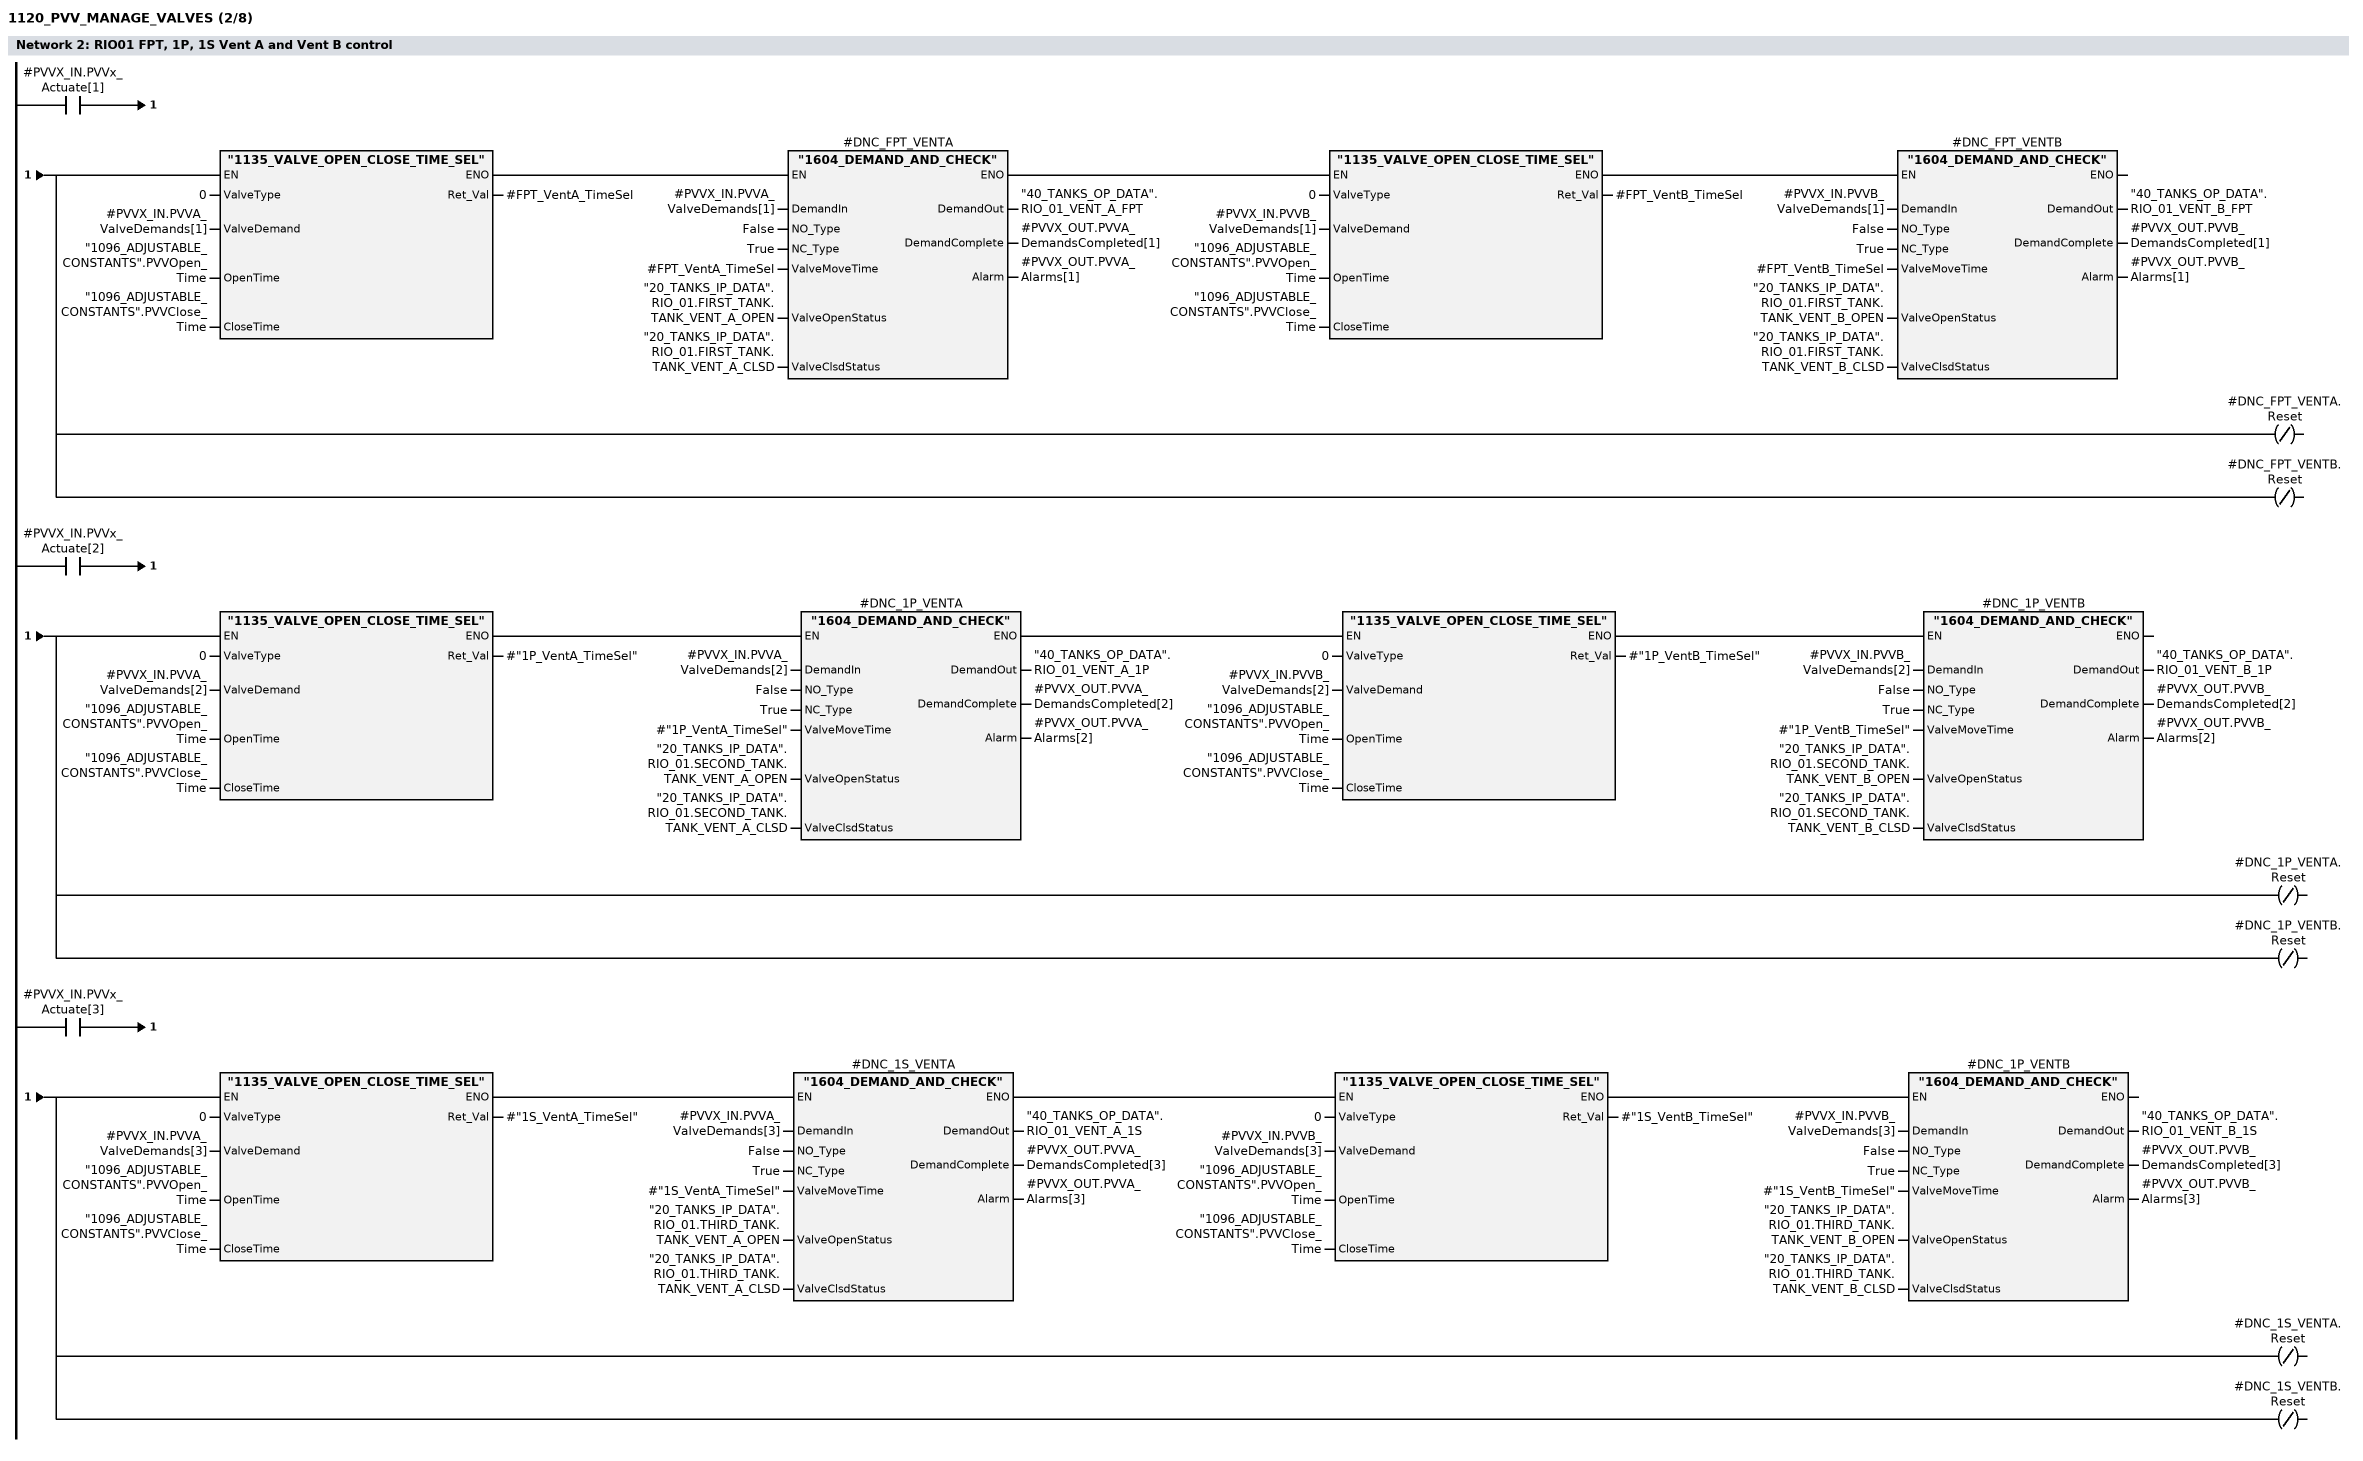
   RUNG wire#powerrail
      Contact( #PVVX_IN.PVVx_Actuate[1] )
      wire#w1
      "1135_VALVE_OPEN_CLOSE_TIME_SEL"(ValveType := 0, ValveDemand := #PVVX_IN.PVVA_ValveDemands[1], OpenTime := "1096_ADJUSTABLE_CONSTANTS".PVVOpen_Time, CloseTime := "1096_ADJUSTABLE_CONSTANTS".PVVClose_Time, Ret_Val => #FPT_VentA_TimeSel)
      #DNC_FPT_VENTA(DemandIn := #PVVX_IN.PVVA_ValveDemands[1], NO_Type := False, NC_Type := True, ValveMoveTime := #FPT_VentA_TimeSel, ValveOpenStatus := "20_TANKS_IP_DATA".RIO_01.FIRST_TANK.TANK_VENT_A_OPEN, ValveClsdStatus := "20_TANKS_IP_DATA".RIO_01.FIRST_TANK.TANK_VENT_A_CLSD, DemandOut => "40_TANKS_OP_DATA".RIO_01_VENT_A_FPT, DemandComplete => #PVVX_OUT.PVVA_DemandsCompleted[1], Alarm => #PVVX_OUT.PVVA_Alarms[1])
      "1135_VALVE_OPEN_CLOSE_TIME_SEL"(ValveType := 0, ValveDemand := #PVVX_IN.PVVB_ValveDemands[1], OpenTime := "1096_ADJUSTABLE_CONSTANTS".PVVOpen_Time, CloseTime := "1096_ADJUSTABLE_CONSTANTS".PVVClose_Time, Ret_Val => #FPT_VentB_TimeSel)
      #DNC_FPT_VENTB(DemandIn := #PVVX_IN.PVVB_ValveDemands[1], NO_Type := False, NC_Type := True, ValveMoveTime := #FPT_VentB_TimeSel, ValveOpenStatus := "20_TANKS_IP_DATA".RIO_01.FIRST_TANK.TANK_VENT_B_OPEN, ValveClsdStatus := "20_TANKS_IP_DATA".RIO_01.FIRST_TANK.TANK_VENT_B_CLSD, DemandOut => "40_TANKS_OP_DATA".RIO_01_VENT_B_FPT, DemandComplete => #PVVX_OUT.PVVB_DemandsCompleted[1], Alarm => #PVVX_OUT.PVVB_Alarms[1])
   END_RUNG
   RUNG wire#w1
      I_Coil( #DNC_FPT_VENTA.Reset )
   END_RUNG
   RUNG wire#w1
      I_Coil( #DNC_FPT_VENTB.Reset )
   END_RUNG
   RUNG wire#powerrail
      Contact( #PVVX_IN.PVVx_Actuate[2] )
      wire#w2
      "1135_VALVE_OPEN_CLOSE_TIME_SEL"(ValveType := 0, ValveDemand := #PVVX_IN.PVVA_ValveDemands[2], OpenTime := "1096_ADJUSTABLE_CONSTANTS".PVVOpen_Time, CloseTime := "1096_ADJUSTABLE_CONSTANTS".PVVClose_Time, Ret_Val => #"1P_VentA_TimeSel")
      #DNC_1P_VENTA(DemandIn := #PVVX_IN.PVVA_ValveDemands[2], NO_Type := False, NC_Type := True, ValveMoveTime := #"1P_VentA_TimeSel", ValveOpenStatus := "20_TANKS_IP_DATA".RIO_01.SECOND_TANK.TANK_VENT_A_OPEN, ValveClsdStatus := "20_TANKS_IP_DATA".RIO_01.SECOND_TANK.TANK_VENT_A_CLSD, DemandOut => "40_TANKS_OP_DATA".RIO_01_VENT_A_1P, DemandComplete => #PVVX_OUT.PVVA_DemandsCompleted[2], Alarm => #PVVX_OUT.PVVA_Alarms[2])
      "1135_VALVE_OPEN_CLOSE_TIME_SEL"(ValveType := 0, ValveDemand := #PVVX_IN.PVVB_ValveDemands[2], OpenTime := "1096_ADJUSTABLE_CONSTANTS".PVVOpen_Time, CloseTime := "1096_ADJUSTABLE_CONSTANTS".PVVClose_Time, Ret_Val => #"1P_VentB_TimeSel")
      #DNC_1P_VENTB(DemandIn := #PVVX_IN.PVVB_ValveDemands[2], NO_Type := False, NC_Type := True, ValveMoveTime := #"1P_VentB_TimeSel", ValveOpenStatus := "20_TANKS_IP_DATA".RIO_01.SECOND_TANK.TANK_VENT_B_OPEN, ValveClsdStatus := "20_TANKS_IP_DATA".RIO_01.SECOND_TANK.TANK_VENT_B_CLSD, DemandOut => "40_TANKS_OP_DATA".RIO_01_VENT_B_1P, DemandComplete => #PVVX_OUT.PVVB_DemandsCompleted[2], Alarm => #PVVX_OUT.PVVB_Alarms[2])
   END_RUNG
   RUNG wire#w2
      I_Coil( #DNC_1P_VENTA.Reset )
   END_RUNG
   RUNG wire#w2
      I_Coil( #DNC_1P_VENTB.Reset )
   END_RUNG
   RUNG wire#powerrail
      Contact( #PVVX_IN.PVVx_Actuate[3] )
      wire#w3
      "1135_VALVE_OPEN_CLOSE_TIME_SEL"(ValveType := 0, ValveDemand := #PVVX_IN.PVVA_ValveDemands[3], OpenTime := "1096_ADJUSTABLE_CONSTANTS".PVVOpen_Time, CloseTime := "1096_ADJUSTABLE_CONSTANTS".PVVClose_Time, Ret_Val => #"1S_VentA_TimeSel")
      #DNC_1S_VENTA(DemandIn := #PVVX_IN.PVVA_ValveDemands[3], NO_Type := False, NC_Type := True, ValveMoveTime := #"1S_VentA_TimeSel", ValveOpenStatus := "20_TANKS_IP_DATA".RIO_01.THIRD_TANK.TANK_VENT_A_OPEN, ValveClsdStatus := "20_TANKS_IP_DATA".RIO_01.THIRD_TANK.TANK_VENT_A_CLSD, DemandOut => "40_TANKS_OP_DATA".RIO_01_VENT_A_1S, DemandComplete => #PVVX_OUT.PVVA_DemandsCompleted[3], Alarm => #PVVX_OUT.PVVA_Alarms[3])
      "1135_VALVE_OPEN_CLOSE_TIME_SEL"(ValveType := 0, ValveDemand := #PVVX_IN.PVVB_ValveDemands[3], OpenTime := "1096_ADJUSTABLE_CONSTANTS".PVVOpen_Time, CloseTime := "1096_ADJUSTABLE_CONSTANTS".PVVClose_Time, Ret_Val => #"1S_VentB_TimeSel")
      #DNC_1P_VENTB(DemandIn := #PVVX_IN.PVVB_ValveDemands[3], NO_Type := False, NC_Type := True, ValveMoveTime := #"1S_VentB_TimeSel", ValveOpenStatus := "20_TANKS_IP_DATA".RIO_01.THIRD_TANK.TANK_VENT_B_OPEN, ValveClsdStatus := "20_TANKS_IP_DATA".RIO_01.THIRD_TANK.TANK_VENT_B_CLSD, DemandOut => "40_TANKS_OP_DATA".RIO_01_VENT_B_1S, DemandComplete => #PVVX_OUT.PVVB_DemandsCompleted[3], Alarm => #PVVX_OUT.PVVB_Alarms[3])
   END_RUNG
   RUNG wire#w3
      I_Coil( #DNC_1S_VENTA.Reset )
   END_RUNG
   RUNG wire#w3
      I_Coil( #DNC_1S_VENTB.Reset )
   END_RUNG
   // the same network as SCL:
   #FPT_VentA_TimeSel := "1135_VALVE_OPEN_CLOSE_TIME_SEL"(EN := #PVVX_IN.PVVx_Actuate[1],
                           ValveType := 0,
                           ValveDemand := #PVVX_IN.PVVA_ValveDemands[1],
                           OpenTime := "1096_ADJUSTABLE_CONSTANTS".PVVOpen_Time,
                           CloseTime := "1096_ADJUSTABLE_CONSTANTS".PVVClose_Time,
                           ENO => #_w1);
   #DNC_FPT_VENTA(EN := #_w1,   // "1604_DEMAND_AND_CHECK"
                  DemandIn := #PVVX_IN.PVVA_ValveDemands[1],
                  NO_Type := False,
                  NC_Type := True,
                  ValveMoveTime := #FPT_VentA_TimeSel,
                  ValveOpenStatus := "20_TANKS_IP_DATA".RIO_01.FIRST_TANK.TANK_VENT_A_OPEN,
                  ValveClsdStatus := "20_TANKS_IP_DATA".RIO_01.FIRST_TANK.TANK_VENT_A_CLSD,
                  DemandOut => "40_TANKS_OP_DATA".RIO_01_VENT_A_FPT,
                  DemandComplete => #PVVX_OUT.PVVA_DemandsCompleted[1],
                  Alarm => #PVVX_OUT.PVVA_Alarms[1],
                  ENO => #_w2);
   #FPT_VentB_TimeSel := "1135_VALVE_OPEN_CLOSE_TIME_SEL"(EN := #_w2,
                           ValveType := 0,
                           ValveDemand := #PVVX_IN.PVVB_ValveDemands[1],
                           OpenTime := "1096_ADJUSTABLE_CONSTANTS".PVVOpen_Time,
                           CloseTime := "1096_ADJUSTABLE_CONSTANTS".PVVClose_Time,
                           ENO => #_w3);
   IF #_w3 THEN
       #DNC_FPT_VENTB(DemandIn := #PVVX_IN.PVVB_ValveDemands[1],   // "1604_DEMAND_AND_CHECK"
                      NO_Type := False,
                      NC_Type := True,
                      ValveMoveTime := #FPT_VentB_TimeSel,
                      ValveOpenStatus := "20_TANKS_IP_DATA".RIO_01.FIRST_TANK.TANK_VENT_B_OPEN,
                      ValveClsdStatus := "20_TANKS_IP_DATA".RIO_01.FIRST_TANK.TANK_VENT_B_CLSD,
                      DemandOut => "40_TANKS_OP_DATA".RIO_01_VENT_B_FPT,
                      DemandComplete => #PVVX_OUT.PVVB_DemandsCompleted[1],
                      Alarm => #PVVX_OUT.PVVB_Alarms[1]);
   END_IF;
   #DNC_FPT_VENTA.Reset := NOT #PVVX_IN.PVVx_Actuate[1];
   #DNC_FPT_VENTB.Reset := NOT #PVVX_IN.PVVx_Actuate[1];
   #"1P_VentA_TimeSel" := "1135_VALVE_OPEN_CLOSE_TIME_SEL"(EN := #PVVX_IN.PVVx_Actuate[2],
                           ValveType := 0,
                           ValveDemand := #PVVX_IN.PVVA_ValveDemands[2],
                           OpenTime := "1096_ADJUSTABLE_CONSTANTS".PVVOpen_Time,
                           CloseTime := "1096_ADJUSTABLE_CONSTANTS".PVVClose_Time,
                           ENO => #_w4);
   #DNC_1P_VENTA(EN := #_w4,   // "1604_DEMAND_AND_CHECK"
                 DemandIn := #PVVX_IN.PVVA_ValveDemands[2],
                 NO_Type := False,
                 NC_Type := True,
                 ValveMoveTime := #"1P_VentA_TimeSel",
                 ValveOpenStatus := "20_TANKS_IP_DATA".RIO_01.SECOND_TANK.TANK_VENT_A_OPEN,
                 ValveClsdStatus := "20_TANKS_IP_DATA".RIO_01.SECOND_TANK.TANK_VENT_A_CLSD,
                 DemandOut => "40_TANKS_OP_DATA".RIO_01_VENT_A_1P,
                 DemandComplete => #PVVX_OUT.PVVA_DemandsCompleted[2],
                 Alarm => #PVVX_OUT.PVVA_Alarms[2],
                 ENO => #_w5);
   #"1P_VentB_TimeSel" := "1135_VALVE_OPEN_CLOSE_TIME_SEL"(EN := #_w5,
                           ValveType := 0,
                           ValveDemand := #PVVX_IN.PVVB_ValveDemands[2],
                           OpenTime := "1096_ADJUSTABLE_CONSTANTS".PVVOpen_Time,
                           CloseTime := "1096_ADJUSTABLE_CONSTANTS".PVVClose_Time,
                           ENO => #_w6);
   IF #_w6 THEN
       #DNC_1P_VENTB(DemandIn := #PVVX_IN.PVVB_ValveDemands[2],   // "1604_DEMAND_AND_CHECK"
                     NO_Type := False,
                     NC_Type := True,
                     ValveMoveTime := #"1P_VentB_TimeSel",
                     ValveOpenStatus := "20_TANKS_IP_DATA".RIO_01.SECOND_TANK.TANK_VENT_B_OPEN,
                     ValveClsdStatus := "20_TANKS_IP_DATA".RIO_01.SECOND_TANK.TANK_VENT_B_CLSD,
                     DemandOut => "40_TANKS_OP_DATA".RIO_01_VENT_B_1P,
                     DemandComplete => #PVVX_OUT.PVVB_DemandsCompleted[2],
                     Alarm => #PVVX_OUT.PVVB_Alarms[2]);
   END_IF;
   #DNC_1P_VENTA.Reset := NOT #PVVX_IN.PVVx_Actuate[2];
   #DNC_1P_VENTB.Reset := NOT #PVVX_IN.PVVx_Actuate[2];
   #"1S_VentA_TimeSel" := "1135_VALVE_OPEN_CLOSE_TIME_SEL"(EN := #PVVX_IN.PVVx_Actuate[3],
                           ValveType := 0,
                           ValveDemand := #PVVX_IN.PVVA_ValveDemands[3],
                           OpenTime := "1096_ADJUSTABLE_CONSTANTS".PVVOpen_Time,
                           CloseTime := "1096_ADJUSTABLE_CONSTANTS".PVVClose_Time,
                           ENO => #_w7);
   #DNC_1S_VENTA(EN := #_w7,   // "1604_DEMAND_AND_CHECK"
                 DemandIn := #PVVX_IN.PVVA_ValveDemands[3],
                 NO_Type := False,
                 NC_Type := True,
                 ValveMoveTime := #"1S_VentA_TimeSel",
                 ValveOpenStatus := "20_TANKS_IP_DATA".RIO_01.THIRD_TANK.TANK_VENT_A_OPEN,
                 ValveClsdStatus := "20_TANKS_IP_DATA".RIO_01.THIRD_TANK.TANK_VENT_A_CLSD,
                 DemandOut => "40_TANKS_OP_DATA".RIO_01_VENT_A_1S,
                 DemandComplete => #PVVX_OUT.PVVA_DemandsCompleted[3],
                 Alarm => #PVVX_OUT.PVVA_Alarms[3],
                 ENO => #_w8);
   #"1S_VentB_TimeSel" := "1135_VALVE_OPEN_CLOSE_TIME_SEL"(EN := #_w8,
                           ValveType := 0,
                           ValveDemand := #PVVX_IN.PVVB_ValveDemands[3],
                           OpenTime := "1096_ADJUSTABLE_CONSTANTS".PVVOpen_Time,
                           CloseTime := "1096_ADJUSTABLE_CONSTANTS".PVVClose_Time,
                           ENO => #_w9);
   IF #_w9 THEN
       #DNC_1P_VENTB(DemandIn := #PVVX_IN.PVVB_ValveDemands[3],   // "1604_DEMAND_AND_CHECK"
                     NO_Type := False,
                     NC_Type := True,
                     ValveMoveTime := #"1S_VentB_TimeSel",
                     ValveOpenStatus := "20_TANKS_IP_DATA".RIO_01.THIRD_TANK.TANK_VENT_B_OPEN,
                     ValveClsdStatus := "20_TANKS_IP_DATA".RIO_01.THIRD_TANK.TANK_VENT_B_CLSD,
                     DemandOut => "40_TANKS_OP_DATA".RIO_01_VENT_B_1S,
                     DemandComplete => #PVVX_OUT.PVVB_DemandsCompleted[3],
                     Alarm => #PVVX_OUT.PVVB_Alarms[3]);
   END_IF;
   #DNC_1S_VENTA.Reset := NOT #PVVX_IN.PVVx_Actuate[3];
   #DNC_1S_VENTB.Reset := NOT #PVVX_IN.PVVx_Actuate[3];
END_REGION

REGION Network 3: RIO02 2P, 2S Vent A and Vent B control
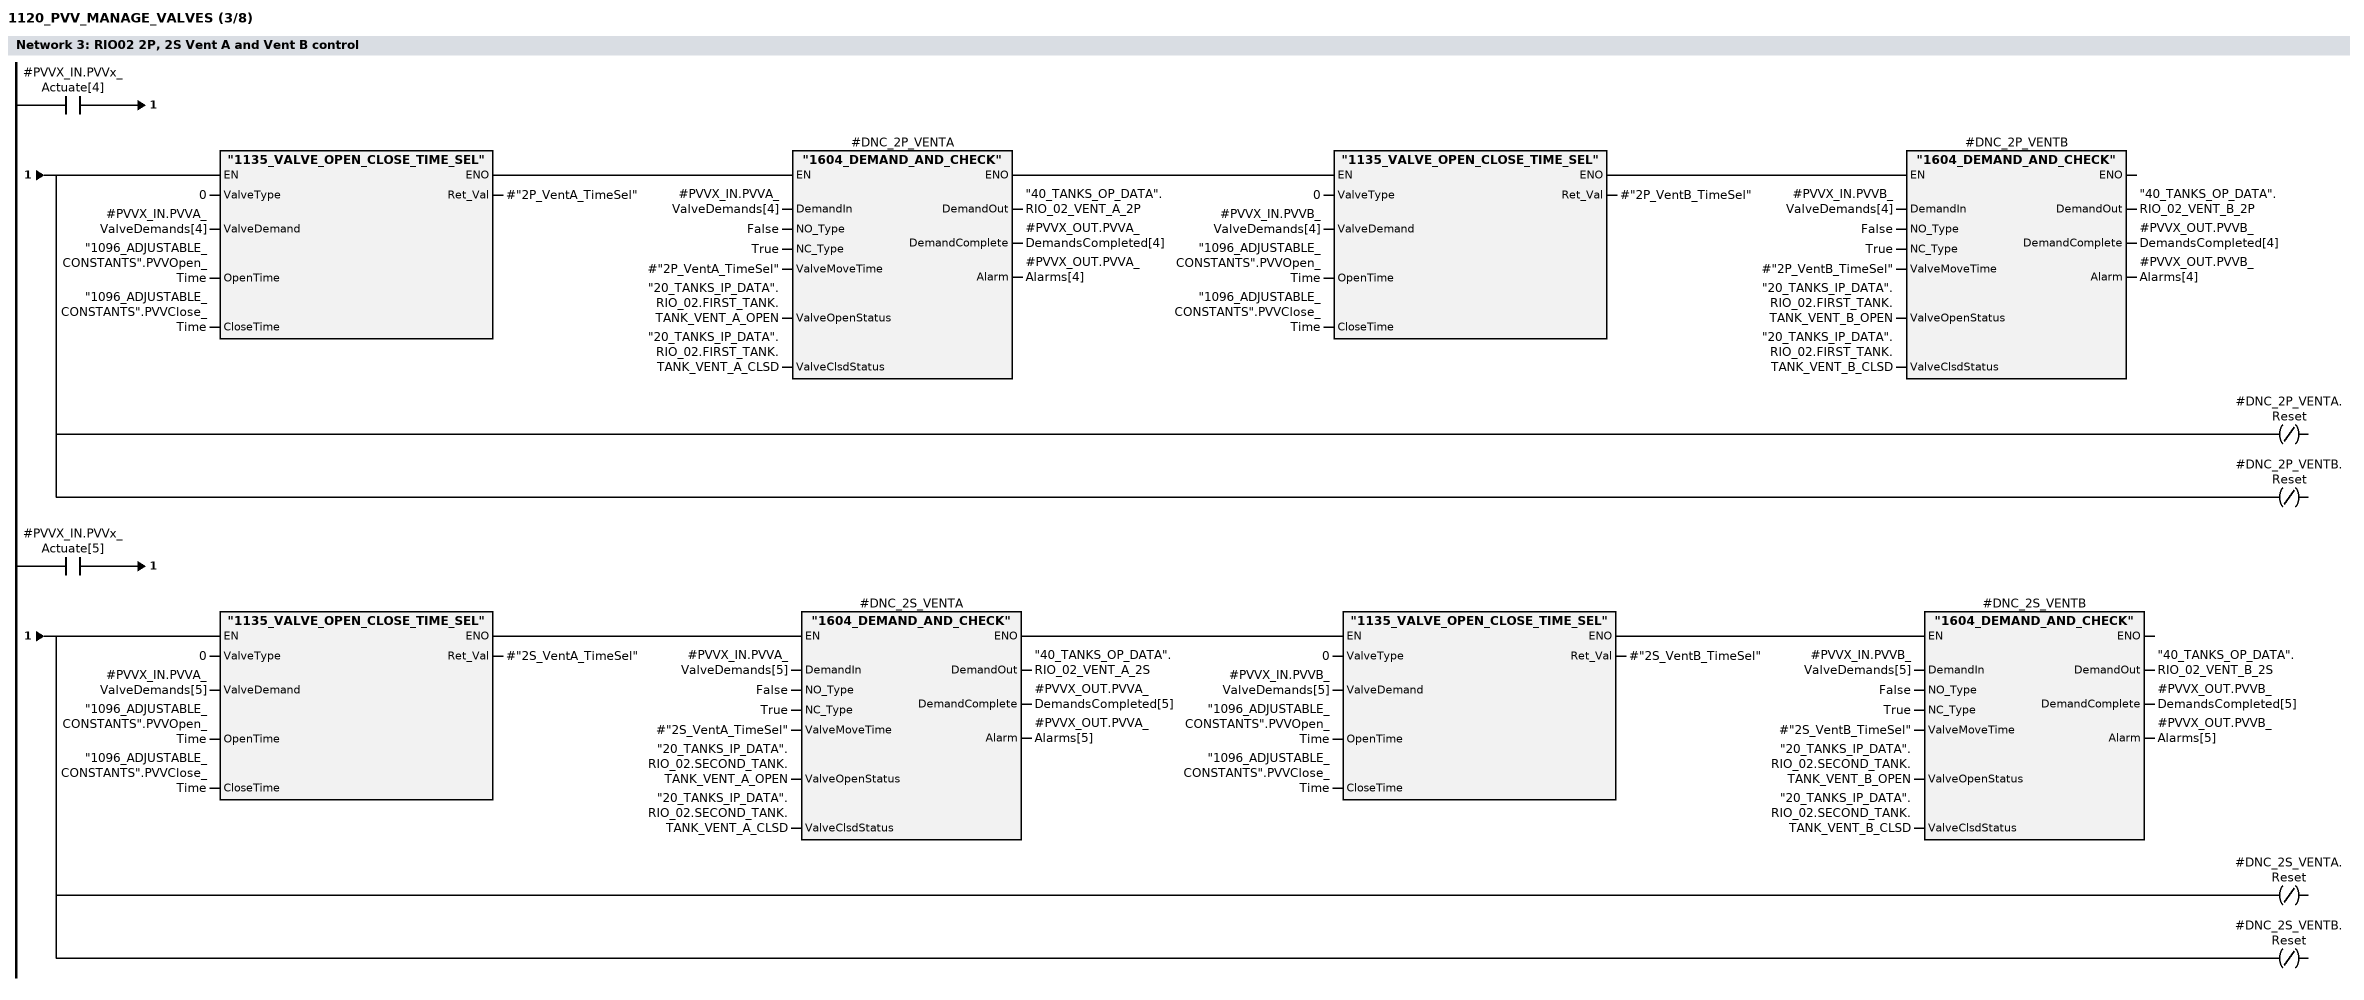
   RUNG wire#powerrail
      Contact( #PVVX_IN.PVVx_Actuate[4] )
      wire#w1
      "1135_VALVE_OPEN_CLOSE_TIME_SEL"(ValveType := 0, ValveDemand := #PVVX_IN.PVVA_ValveDemands[4], OpenTime := "1096_ADJUSTABLE_CONSTANTS".PVVOpen_Time, CloseTime := "1096_ADJUSTABLE_CONSTANTS".PVVClose_Time, Ret_Val => #"2P_VentA_TimeSel")
      #DNC_2P_VENTA(DemandIn := #PVVX_IN.PVVA_ValveDemands[4], NO_Type := False, NC_Type := True, ValveMoveTime := #"2P_VentA_TimeSel", ValveOpenStatus := "20_TANKS_IP_DATA".RIO_02.FIRST_TANK.TANK_VENT_A_OPEN, ValveClsdStatus := "20_TANKS_IP_DATA".RIO_02.FIRST_TANK.TANK_VENT_A_CLSD, DemandOut => "40_TANKS_OP_DATA".RIO_02_VENT_A_2P, DemandComplete => #PVVX_OUT.PVVA_DemandsCompleted[4], Alarm => #PVVX_OUT.PVVA_Alarms[4])
      "1135_VALVE_OPEN_CLOSE_TIME_SEL"(ValveType := 0, ValveDemand := #PVVX_IN.PVVB_ValveDemands[4], OpenTime := "1096_ADJUSTABLE_CONSTANTS".PVVOpen_Time, CloseTime := "1096_ADJUSTABLE_CONSTANTS".PVVClose_Time, Ret_Val => #"2P_VentB_TimeSel")
      #DNC_2P_VENTB(DemandIn := #PVVX_IN.PVVB_ValveDemands[4], NO_Type := False, NC_Type := True, ValveMoveTime := #"2P_VentB_TimeSel", ValveOpenStatus := "20_TANKS_IP_DATA".RIO_02.FIRST_TANK.TANK_VENT_B_OPEN, ValveClsdStatus := "20_TANKS_IP_DATA".RIO_02.FIRST_TANK.TANK_VENT_B_CLSD, DemandOut => "40_TANKS_OP_DATA".RIO_02_VENT_B_2P, DemandComplete => #PVVX_OUT.PVVB_DemandsCompleted[4], Alarm => #PVVX_OUT.PVVB_Alarms[4])
   END_RUNG
   RUNG wire#w1
      I_Coil( #DNC_2P_VENTA.Reset )
   END_RUNG
   RUNG wire#w1
      I_Coil( #DNC_2P_VENTB.Reset )
   END_RUNG
   RUNG wire#powerrail
      Contact( #PVVX_IN.PVVx_Actuate[5] )
      wire#w2
      "1135_VALVE_OPEN_CLOSE_TIME_SEL"(ValveType := 0, ValveDemand := #PVVX_IN.PVVA_ValveDemands[5], OpenTime := "1096_ADJUSTABLE_CONSTANTS".PVVOpen_Time, CloseTime := "1096_ADJUSTABLE_CONSTANTS".PVVClose_Time, Ret_Val => #"2S_VentA_TimeSel")
      #DNC_2S_VENTA(DemandIn := #PVVX_IN.PVVA_ValveDemands[5], NO_Type := False, NC_Type := True, ValveMoveTime := #"2S_VentA_TimeSel", ValveOpenStatus := "20_TANKS_IP_DATA".RIO_02.SECOND_TANK.TANK_VENT_A_OPEN, ValveClsdStatus := "20_TANKS_IP_DATA".RIO_02.SECOND_TANK.TANK_VENT_A_CLSD, DemandOut => "40_TANKS_OP_DATA".RIO_02_VENT_A_2S, DemandComplete => #PVVX_OUT.PVVA_DemandsCompleted[5], Alarm => #PVVX_OUT.PVVA_Alarms[5])
      "1135_VALVE_OPEN_CLOSE_TIME_SEL"(ValveType := 0, ValveDemand := #PVVX_IN.PVVB_ValveDemands[5], OpenTime := "1096_ADJUSTABLE_CONSTANTS".PVVOpen_Time, CloseTime := "1096_ADJUSTABLE_CONSTANTS".PVVClose_Time, Ret_Val => #"2S_VentB_TimeSel")
      #DNC_2S_VENTB(DemandIn := #PVVX_IN.PVVB_ValveDemands[5], NO_Type := False, NC_Type := True, ValveMoveTime := #"2S_VentB_TimeSel", ValveOpenStatus := "20_TANKS_IP_DATA".RIO_02.SECOND_TANK.TANK_VENT_B_OPEN, ValveClsdStatus := "20_TANKS_IP_DATA".RIO_02.SECOND_TANK.TANK_VENT_B_CLSD, DemandOut => "40_TANKS_OP_DATA".RIO_02_VENT_B_2S, DemandComplete => #PVVX_OUT.PVVB_DemandsCompleted[5], Alarm => #PVVX_OUT.PVVB_Alarms[5])
   END_RUNG
   RUNG wire#w2
      I_Coil( #DNC_2S_VENTA.Reset )
   END_RUNG
   RUNG wire#w2
      I_Coil( #DNC_2S_VENTB.Reset )
   END_RUNG
   // the same network as SCL:
   #"2P_VentA_TimeSel" := "1135_VALVE_OPEN_CLOSE_TIME_SEL"(EN := #PVVX_IN.PVVx_Actuate[4],
                           ValveType := 0,
                           ValveDemand := #PVVX_IN.PVVA_ValveDemands[4],
                           OpenTime := "1096_ADJUSTABLE_CONSTANTS".PVVOpen_Time,
                           CloseTime := "1096_ADJUSTABLE_CONSTANTS".PVVClose_Time,
                           ENO => #_w1);
   #DNC_2P_VENTA(EN := #_w1,   // "1604_DEMAND_AND_CHECK"
                 DemandIn := #PVVX_IN.PVVA_ValveDemands[4],
                 NO_Type := False,
                 NC_Type := True,
                 ValveMoveTime := #"2P_VentA_TimeSel",
                 ValveOpenStatus := "20_TANKS_IP_DATA".RIO_02.FIRST_TANK.TANK_VENT_A_OPEN,
                 ValveClsdStatus := "20_TANKS_IP_DATA".RIO_02.FIRST_TANK.TANK_VENT_A_CLSD,
                 DemandOut => "40_TANKS_OP_DATA".RIO_02_VENT_A_2P,
                 DemandComplete => #PVVX_OUT.PVVA_DemandsCompleted[4],
                 Alarm => #PVVX_OUT.PVVA_Alarms[4],
                 ENO => #_w2);
   #"2P_VentB_TimeSel" := "1135_VALVE_OPEN_CLOSE_TIME_SEL"(EN := #_w2,
                           ValveType := 0,
                           ValveDemand := #PVVX_IN.PVVB_ValveDemands[4],
                           OpenTime := "1096_ADJUSTABLE_CONSTANTS".PVVOpen_Time,
                           CloseTime := "1096_ADJUSTABLE_CONSTANTS".PVVClose_Time,
                           ENO => #_w3);
   IF #_w3 THEN
       #DNC_2P_VENTB(DemandIn := #PVVX_IN.PVVB_ValveDemands[4],   // "1604_DEMAND_AND_CHECK"
                     NO_Type := False,
                     NC_Type := True,
                     ValveMoveTime := #"2P_VentB_TimeSel",
                     ValveOpenStatus := "20_TANKS_IP_DATA".RIO_02.FIRST_TANK.TANK_VENT_B_OPEN,
                     ValveClsdStatus := "20_TANKS_IP_DATA".RIO_02.FIRST_TANK.TANK_VENT_B_CLSD,
                     DemandOut => "40_TANKS_OP_DATA".RIO_02_VENT_B_2P,
                     DemandComplete => #PVVX_OUT.PVVB_DemandsCompleted[4],
                     Alarm => #PVVX_OUT.PVVB_Alarms[4]);
   END_IF;
   #DNC_2P_VENTA.Reset := NOT #PVVX_IN.PVVx_Actuate[4];
   #DNC_2P_VENTB.Reset := NOT #PVVX_IN.PVVx_Actuate[4];
   #"2S_VentA_TimeSel" := "1135_VALVE_OPEN_CLOSE_TIME_SEL"(EN := #PVVX_IN.PVVx_Actuate[5],
                           ValveType := 0,
                           ValveDemand := #PVVX_IN.PVVA_ValveDemands[5],
                           OpenTime := "1096_ADJUSTABLE_CONSTANTS".PVVOpen_Time,
                           CloseTime := "1096_ADJUSTABLE_CONSTANTS".PVVClose_Time,
                           ENO => #_w4);
   #DNC_2S_VENTA(EN := #_w4,   // "1604_DEMAND_AND_CHECK"
                 DemandIn := #PVVX_IN.PVVA_ValveDemands[5],
                 NO_Type := False,
                 NC_Type := True,
                 ValveMoveTime := #"2S_VentA_TimeSel",
                 ValveOpenStatus := "20_TANKS_IP_DATA".RIO_02.SECOND_TANK.TANK_VENT_A_OPEN,
                 ValveClsdStatus := "20_TANKS_IP_DATA".RIO_02.SECOND_TANK.TANK_VENT_A_CLSD,
                 DemandOut => "40_TANKS_OP_DATA".RIO_02_VENT_A_2S,
                 DemandComplete => #PVVX_OUT.PVVA_DemandsCompleted[5],
                 Alarm => #PVVX_OUT.PVVA_Alarms[5],
                 ENO => #_w5);
   #"2S_VentB_TimeSel" := "1135_VALVE_OPEN_CLOSE_TIME_SEL"(EN := #_w5,
                           ValveType := 0,
                           ValveDemand := #PVVX_IN.PVVB_ValveDemands[5],
                           OpenTime := "1096_ADJUSTABLE_CONSTANTS".PVVOpen_Time,
                           CloseTime := "1096_ADJUSTABLE_CONSTANTS".PVVClose_Time,
                           ENO => #_w6);
   IF #_w6 THEN
       #DNC_2S_VENTB(DemandIn := #PVVX_IN.PVVB_ValveDemands[5],   // "1604_DEMAND_AND_CHECK"
                     NO_Type := False,
                     NC_Type := True,
                     ValveMoveTime := #"2S_VentB_TimeSel",
                     ValveOpenStatus := "20_TANKS_IP_DATA".RIO_02.SECOND_TANK.TANK_VENT_B_OPEN,
                     ValveClsdStatus := "20_TANKS_IP_DATA".RIO_02.SECOND_TANK.TANK_VENT_B_CLSD,
                     DemandOut => "40_TANKS_OP_DATA".RIO_02_VENT_B_2S,
                     DemandComplete => #PVVX_OUT.PVVB_DemandsCompleted[5],
                     Alarm => #PVVX_OUT.PVVB_Alarms[5]);
   END_IF;
   #DNC_2S_VENTA.Reset := NOT #PVVX_IN.PVVx_Actuate[5];
   #DNC_2S_VENTB.Reset := NOT #PVVX_IN.PVVx_Actuate[5];
END_REGION

REGION Network 4: RIO02 3P, 3S Vent A and Vent B control
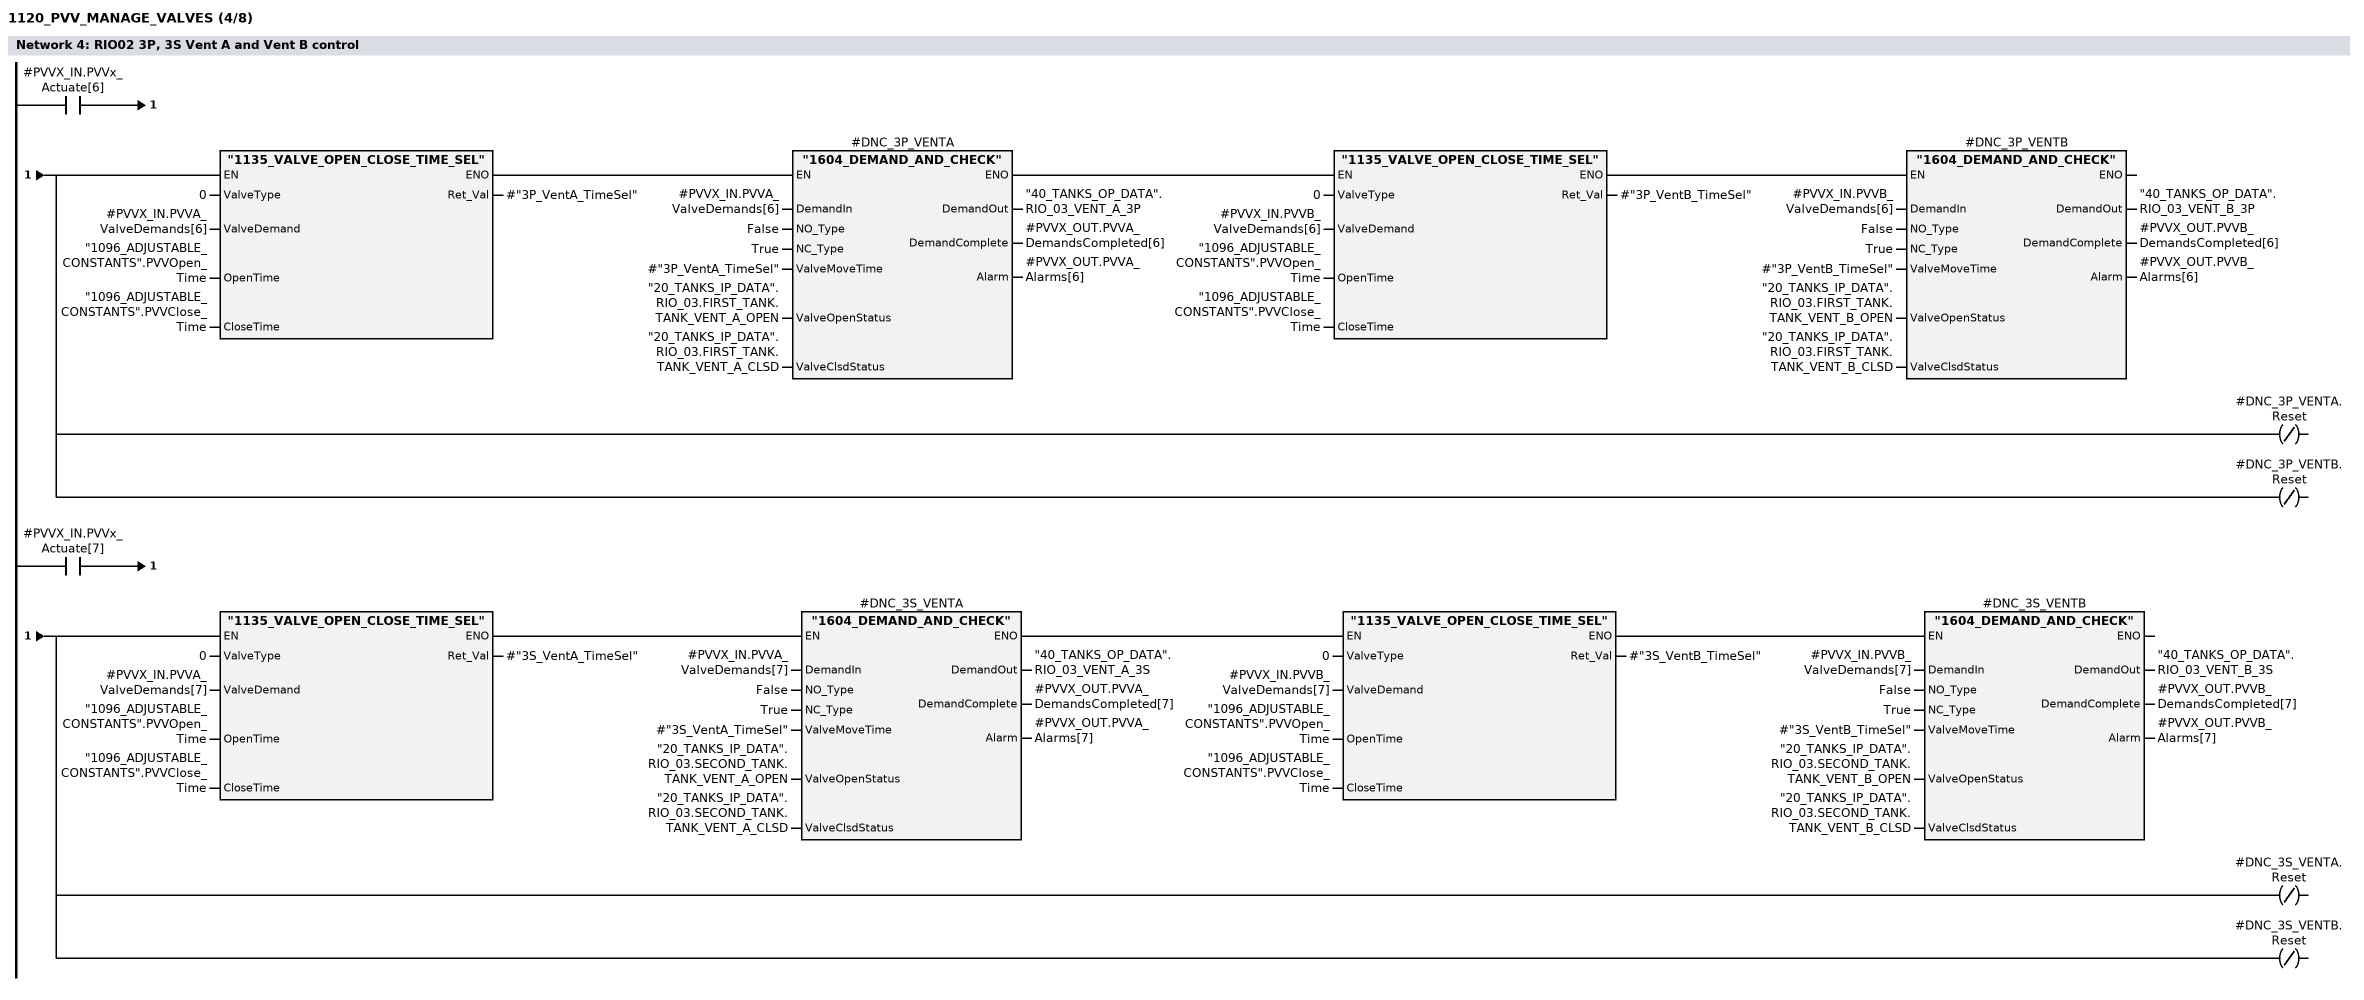
   RUNG wire#powerrail
      Contact( #PVVX_IN.PVVx_Actuate[6] )
      wire#w1
      "1135_VALVE_OPEN_CLOSE_TIME_SEL"(ValveType := 0, ValveDemand := #PVVX_IN.PVVA_ValveDemands[6], OpenTime := "1096_ADJUSTABLE_CONSTANTS".PVVOpen_Time, CloseTime := "1096_ADJUSTABLE_CONSTANTS".PVVClose_Time, Ret_Val => #"3P_VentA_TimeSel")
      #DNC_3P_VENTA(DemandIn := #PVVX_IN.PVVA_ValveDemands[6], NO_Type := False, NC_Type := True, ValveMoveTime := #"3P_VentA_TimeSel", ValveOpenStatus := "20_TANKS_IP_DATA".RIO_03.FIRST_TANK.TANK_VENT_A_OPEN, ValveClsdStatus := "20_TANKS_IP_DATA".RIO_03.FIRST_TANK.TANK_VENT_A_CLSD, DemandOut => "40_TANKS_OP_DATA".RIO_03_VENT_A_3P, DemandComplete => #PVVX_OUT.PVVA_DemandsCompleted[6], Alarm => #PVVX_OUT.PVVA_Alarms[6])
      "1135_VALVE_OPEN_CLOSE_TIME_SEL"(ValveType := 0, ValveDemand := #PVVX_IN.PVVB_ValveDemands[6], OpenTime := "1096_ADJUSTABLE_CONSTANTS".PVVOpen_Time, CloseTime := "1096_ADJUSTABLE_CONSTANTS".PVVClose_Time, Ret_Val => #"3P_VentB_TimeSel")
      #DNC_3P_VENTB(DemandIn := #PVVX_IN.PVVB_ValveDemands[6], NO_Type := False, NC_Type := True, ValveMoveTime := #"3P_VentB_TimeSel", ValveOpenStatus := "20_TANKS_IP_DATA".RIO_03.FIRST_TANK.TANK_VENT_B_OPEN, ValveClsdStatus := "20_TANKS_IP_DATA".RIO_03.FIRST_TANK.TANK_VENT_B_CLSD, DemandOut => "40_TANKS_OP_DATA".RIO_03_VENT_B_3P, DemandComplete => #PVVX_OUT.PVVB_DemandsCompleted[6], Alarm => #PVVX_OUT.PVVB_Alarms[6])
   END_RUNG
   RUNG wire#w1
      I_Coil( #DNC_3P_VENTA.Reset )
   END_RUNG
   RUNG wire#w1
      I_Coil( #DNC_3P_VENTB.Reset )
   END_RUNG
   RUNG wire#powerrail
      Contact( #PVVX_IN.PVVx_Actuate[7] )
      wire#w2
      "1135_VALVE_OPEN_CLOSE_TIME_SEL"(ValveType := 0, ValveDemand := #PVVX_IN.PVVA_ValveDemands[7], OpenTime := "1096_ADJUSTABLE_CONSTANTS".PVVOpen_Time, CloseTime := "1096_ADJUSTABLE_CONSTANTS".PVVClose_Time, Ret_Val => #"3S_VentA_TimeSel")
      #DNC_3S_VENTA(DemandIn := #PVVX_IN.PVVA_ValveDemands[7], NO_Type := False, NC_Type := True, ValveMoveTime := #"3S_VentA_TimeSel", ValveOpenStatus := "20_TANKS_IP_DATA".RIO_03.SECOND_TANK.TANK_VENT_A_OPEN, ValveClsdStatus := "20_TANKS_IP_DATA".RIO_03.SECOND_TANK.TANK_VENT_A_CLSD, DemandOut => "40_TANKS_OP_DATA".RIO_03_VENT_A_3S, DemandComplete => #PVVX_OUT.PVVA_DemandsCompleted[7], Alarm => #PVVX_OUT.PVVA_Alarms[7])
      "1135_VALVE_OPEN_CLOSE_TIME_SEL"(ValveType := 0, ValveDemand := #PVVX_IN.PVVB_ValveDemands[7], OpenTime := "1096_ADJUSTABLE_CONSTANTS".PVVOpen_Time, CloseTime := "1096_ADJUSTABLE_CONSTANTS".PVVClose_Time, Ret_Val => #"3S_VentB_TimeSel")
      #DNC_3S_VENTB(DemandIn := #PVVX_IN.PVVB_ValveDemands[7], NO_Type := False, NC_Type := True, ValveMoveTime := #"3S_VentB_TimeSel", ValveOpenStatus := "20_TANKS_IP_DATA".RIO_03.SECOND_TANK.TANK_VENT_B_OPEN, ValveClsdStatus := "20_TANKS_IP_DATA".RIO_03.SECOND_TANK.TANK_VENT_B_CLSD, DemandOut => "40_TANKS_OP_DATA".RIO_03_VENT_B_3S, DemandComplete => #PVVX_OUT.PVVB_DemandsCompleted[7], Alarm => #PVVX_OUT.PVVB_Alarms[7])
   END_RUNG
   RUNG wire#w2
      I_Coil( #DNC_3S_VENTA.Reset )
   END_RUNG
   RUNG wire#w2
      I_Coil( #DNC_3S_VENTB.Reset )
   END_RUNG
   // the same network as SCL:
   #"3P_VentA_TimeSel" := "1135_VALVE_OPEN_CLOSE_TIME_SEL"(EN := #PVVX_IN.PVVx_Actuate[6],
                           ValveType := 0,
                           ValveDemand := #PVVX_IN.PVVA_ValveDemands[6],
                           OpenTime := "1096_ADJUSTABLE_CONSTANTS".PVVOpen_Time,
                           CloseTime := "1096_ADJUSTABLE_CONSTANTS".PVVClose_Time,
                           ENO => #_w1);
   #DNC_3P_VENTA(EN := #_w1,   // "1604_DEMAND_AND_CHECK"
                 DemandIn := #PVVX_IN.PVVA_ValveDemands[6],
                 NO_Type := False,
                 NC_Type := True,
                 ValveMoveTime := #"3P_VentA_TimeSel",
                 ValveOpenStatus := "20_TANKS_IP_DATA".RIO_03.FIRST_TANK.TANK_VENT_A_OPEN,
                 ValveClsdStatus := "20_TANKS_IP_DATA".RIO_03.FIRST_TANK.TANK_VENT_A_CLSD,
                 DemandOut => "40_TANKS_OP_DATA".RIO_03_VENT_A_3P,
                 DemandComplete => #PVVX_OUT.PVVA_DemandsCompleted[6],
                 Alarm => #PVVX_OUT.PVVA_Alarms[6],
                 ENO => #_w2);
   #"3P_VentB_TimeSel" := "1135_VALVE_OPEN_CLOSE_TIME_SEL"(EN := #_w2,
                           ValveType := 0,
                           ValveDemand := #PVVX_IN.PVVB_ValveDemands[6],
                           OpenTime := "1096_ADJUSTABLE_CONSTANTS".PVVOpen_Time,
                           CloseTime := "1096_ADJUSTABLE_CONSTANTS".PVVClose_Time,
                           ENO => #_w3);
   IF #_w3 THEN
       #DNC_3P_VENTB(DemandIn := #PVVX_IN.PVVB_ValveDemands[6],   // "1604_DEMAND_AND_CHECK"
                     NO_Type := False,
                     NC_Type := True,
                     ValveMoveTime := #"3P_VentB_TimeSel",
                     ValveOpenStatus := "20_TANKS_IP_DATA".RIO_03.FIRST_TANK.TANK_VENT_B_OPEN,
                     ValveClsdStatus := "20_TANKS_IP_DATA".RIO_03.FIRST_TANK.TANK_VENT_B_CLSD,
                     DemandOut => "40_TANKS_OP_DATA".RIO_03_VENT_B_3P,
                     DemandComplete => #PVVX_OUT.PVVB_DemandsCompleted[6],
                     Alarm => #PVVX_OUT.PVVB_Alarms[6]);
   END_IF;
   #DNC_3P_VENTA.Reset := NOT #PVVX_IN.PVVx_Actuate[6];
   #DNC_3P_VENTB.Reset := NOT #PVVX_IN.PVVx_Actuate[6];
   #"3S_VentA_TimeSel" := "1135_VALVE_OPEN_CLOSE_TIME_SEL"(EN := #PVVX_IN.PVVx_Actuate[7],
                           ValveType := 0,
                           ValveDemand := #PVVX_IN.PVVA_ValveDemands[7],
                           OpenTime := "1096_ADJUSTABLE_CONSTANTS".PVVOpen_Time,
                           CloseTime := "1096_ADJUSTABLE_CONSTANTS".PVVClose_Time,
                           ENO => #_w4);
   #DNC_3S_VENTA(EN := #_w4,   // "1604_DEMAND_AND_CHECK"
                 DemandIn := #PVVX_IN.PVVA_ValveDemands[7],
                 NO_Type := False,
                 NC_Type := True,
                 ValveMoveTime := #"3S_VentA_TimeSel",
                 ValveOpenStatus := "20_TANKS_IP_DATA".RIO_03.SECOND_TANK.TANK_VENT_A_OPEN,
                 ValveClsdStatus := "20_TANKS_IP_DATA".RIO_03.SECOND_TANK.TANK_VENT_A_CLSD,
                 DemandOut => "40_TANKS_OP_DATA".RIO_03_VENT_A_3S,
                 DemandComplete => #PVVX_OUT.PVVA_DemandsCompleted[7],
                 Alarm => #PVVX_OUT.PVVA_Alarms[7],
                 ENO => #_w5);
   #"3S_VentB_TimeSel" := "1135_VALVE_OPEN_CLOSE_TIME_SEL"(EN := #_w5,
                           ValveType := 0,
                           ValveDemand := #PVVX_IN.PVVB_ValveDemands[7],
                           OpenTime := "1096_ADJUSTABLE_CONSTANTS".PVVOpen_Time,
                           CloseTime := "1096_ADJUSTABLE_CONSTANTS".PVVClose_Time,
                           ENO => #_w6);
   IF #_w6 THEN
       #DNC_3S_VENTB(DemandIn := #PVVX_IN.PVVB_ValveDemands[7],   // "1604_DEMAND_AND_CHECK"
                     NO_Type := False,
                     NC_Type := True,
                     ValveMoveTime := #"3S_VentB_TimeSel",
                     ValveOpenStatus := "20_TANKS_IP_DATA".RIO_03.SECOND_TANK.TANK_VENT_B_OPEN,
                     ValveClsdStatus := "20_TANKS_IP_DATA".RIO_03.SECOND_TANK.TANK_VENT_B_CLSD,
                     DemandOut => "40_TANKS_OP_DATA".RIO_03_VENT_B_3S,
                     DemandComplete => #PVVX_OUT.PVVB_DemandsCompleted[7],
                     Alarm => #PVVX_OUT.PVVB_Alarms[7]);
   END_IF;
   #DNC_3S_VENTA.Reset := NOT #PVVX_IN.PVVx_Actuate[7];
   #DNC_3S_VENTB.Reset := NOT #PVVX_IN.PVVx_Actuate[7];
END_REGION

